(* Logix 5000 project; controller FV vendor 1 type 14 code 217 rev 31.11; software revision 31.00; part 40 of 63 *)
(* tags used below, declared in another part *)
   FV_ALARM : PlantItem;   // ALARM
   FV_ALARM_RawOutput : ALIAS FOR Remote_IO:4:O.Data.5;   // FV_ALARM Audible alarm
   FV_B22 : INT[255];   // YSVFILL_FL YSV filling process flags
   FV_FV25C : PlantItem;   // FV25C
   FV_FV25C_RawOutput : ALIAS FOR Remote_IO:4:O.Data.0;   // FV_FV25C FV 25 cone cooling valve
   FV_FV25J : PlantItem;   // FV25J
   FV_FV25J_RawOutput : ALIAS FOR Remote_IO:4:O.Data.1;   // FV_FV25J FV 25 jacket cooling valve
   FV_FV26C : PlantItem;   // FV26C
   FV_FV26C_RawOutput : ALIAS FOR Remote_IO:9:O.Data.1;   // FV_FV26C FV26 coolant SOV (Cone)
   FV_FV26J : PlantItem;   // FV26J
   FV_FV26J_RawOutput : ALIAS FOR Remote_IO:9:O.Data.0;   // FV_FV26J FV26 coolant SOV (Tank)
   FV_FV27C : PlantItem;   // FV27C
   FV_FV27C_RawOutput : ALIAS FOR Remote_IO:9:O.Data.3;   // FV_FV27C FV27 coolant SOV (Cone)
   FV_FV27J : PlantItem;   // FV27J
   FV_FV27J_RawOutput : ALIAS FOR Remote_IO:9:O.Data.2;   // FV_FV27J FV27 coolant SOV (Tank)
   FV_FV28C : PlantItem;   // FV28C
   FV_FV28C_RawOutput : ALIAS FOR Remote_IO:9:O.Data.5;   // FV_FV28C FV28 coolant SOV (Cone)
   FV_FV28J : PlantItem;   // FV28J
   FV_FV28J_RawOutput : ALIAS FOR Remote_IO:9:O.Data.4;   // FV_FV28J FV28 coolant SOV (Tank)
   FV_FV29C : PlantItem;   // FV29C
   FV_FV29C_RawOutput : ALIAS FOR Remote_IO:9:O.Data.7;   // FV_FV29C FV29 coolant SOV (Cone)
   FV_FV29J : PlantItem;   // FV29J
   FV_FV29J_RawOutput : ALIAS FOR Remote_IO:9:O.Data.6;   // FV_FV29J FV29 coolant SOV (Tank)
   FV_FV30C : PlantItem;   // FV30C
   FV_FV30C_RawOutput : ALIAS FOR Remote_IO:9:O.Data.9;   // FV_FV30C FV30 coolant SOV (Cone)
   FV_FV30J : PlantItem;   // FV30J
   FV_FV30J_RawOutput : ALIAS FOR Remote_IO:9:O.Data.8;   // FV_FV30J FV30 coolant SOV (Tank)
   FV_FV31C : PlantItem;   // FV31C
   FV_FV31C_RawOutput : ALIAS FOR Remote_IO:9:O.Data.11;   // FV_FV31C FV31 coolant SOV (Cone)
   FV_FV31J : PlantItem;   // FV31J
   FV_FV31J_RawOutput : ALIAS FOR Remote_IO:9:O.Data.10;   // FV_FV31J FV31 coolant SOV (Tank)
   FV_N141 : INT[255];   // YSV1 DATA
   FV_N142 : INT[255];   // YSV2 DATA
   FV_N143 : INT[255];   // YSV3 DATA
   FV_N20 : INT[255];   // YSVFILL<PC YSV Filling data fro m PC
   FV_N21 : INT[255];   // YSVFILL>PC YSV Filling process data to PC and contr ol regs
   FV_PUMP1 : PlantItem;   // PUMP1
   FV_PUMP1_RawOutput : ALIAS FOR Remote_IO:4:O.Data.13;   // FV_PUMP1 Coolant recirc.valve 1
   FV_PUMP2 : PlantItem;   // PUMP2
   FV_PUMP2_RawOutput : ALIAS FOR Remote_IO:4:O.Data.14;   // FV_PUMP2 Coolant recirc.valve 2
   FV_PUMP3 : PlantItem;   // PUMP3
   FV_PUMP3_RawOutput : ALIAS FOR Remote_IO:4:O.Data.15;   // FV_PUMP3 Coolant recirc.valve 3
   FV_SOV1 : PlantItem;   // SOV1
   FV_SOV1_RawOutput : ALIAS FOR Remote_IO:5:O.Data.6;   // FV_SOV1 Air supply to reseed pump
   FV_SOV2 : PlantItem;   // SOV2
   FV_SOV2_RawOutput : ALIAS FOR Remote_IO:5:O.Data.7;   // FV_SOV2 Air supply to reseed pump
   FV_T23 : TIMER[10];
   FV_YSV1CV : PlantItem;   // YSV1CV
   FV_YSV1CV_RawOutput : ALIAS FOR Remote_IO:5:O.Data.12;   // FV_YSV1CV
   FV_YSV1J : PlantItem;   // YSV1J
   FV_YSV1J_RawOutput : ALIAS FOR Remote_IO:4:O.Data.9;   // FV_YSV1J YSV 1 cooling valve
   FV_YSV2CV : PlantItem;   // YSV2CV
   FV_YSV2CV_RawOutput : ALIAS FOR Remote_IO:5:O.Data.13;   // FV_YSV2CV
   FV_YSV2J : PlantItem;   // YSV2J
   FV_YSV2J_RawOutput : ALIAS FOR Remote_IO:4:O.Data.11;   // FV_YSV2J YSV 2 cooling valve
   FV_YSV2O : PlantItem;   // YSV2O
   FV_YSV2O_RawOutput : ALIAS FOR Remote_IO:4:O.Data.4;   // FV_YSV2O YSV 2 outlet valve
   FV_YSV2R : PlantItem;   // YSV2R
   FV_YSV2R_RawOutput : ALIAS FOR Remote_IO:4:O.Data.12;   // FV_YSV2R YSV 2 rouser
   FV_YSV3J : PlantItem;   // YSV3J
   FV_YSV3J_RawOutput : ALIAS FOR Remote_IO:4:O.Data.7;   // FV_YSV3J YSV 3 cooling valve
   FV_YSV3O : PlantItem;   // YSV3O
   FV_YSV3O_RawOutput : ALIAS FOR Remote_IO:4:O.Data.6;   // FV_YSV3O YSV 3 outlet valve
   FV_YSV3R : PlantItem;   // YSV3R
   FV_YSV3R_RawOutput : ALIAS FOR Remote_IO:4:O.Data.8;   // FV_YSV3R YSV 3 rouser
(* FV_Common, continued *)

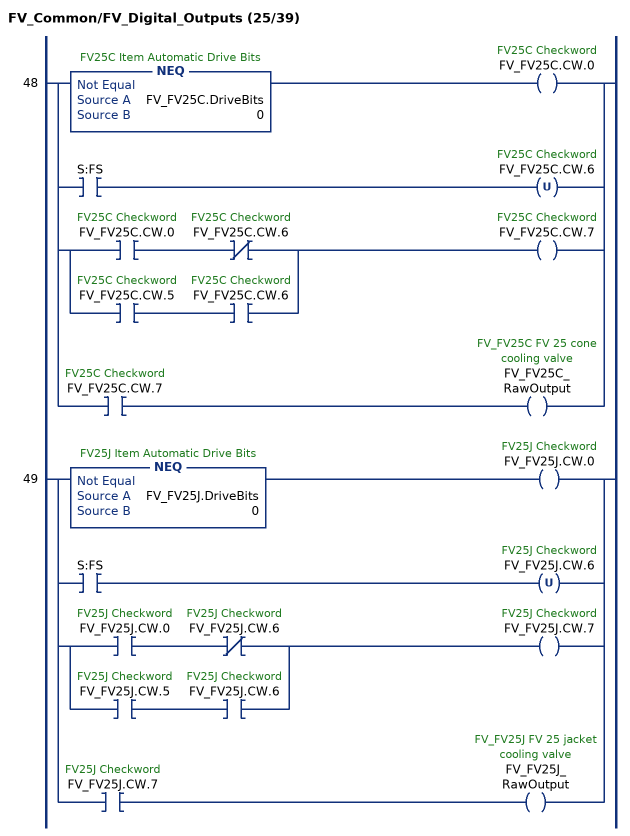
   [picture p849: FV_Common/FV_Digital_Outputs rungs 48-49]
   48: [NEQ(FV_FV25C.DriveBits,0) OTE(FV_FV25C.CW.0) ,XIC(S:FS) OTU(FV_FV25C.CW.6) ,[XIC(FV_FV25C.CW.0) XIO(FV_FV25C.CW.6) ,XIC(FV_FV25C.CW.5) XIC(FV_FV25C.CW.6) ] OTE(FV_FV25C.CW.7) ,XIC(FV_FV25C.CW.7) OTE(FV_FV25C_RawOutput) ];
   49: [NEQ(FV_FV25J.DriveBits,0) OTE(FV_FV25J.CW.0) ,XIC(S:FS) OTU(FV_FV25J.CW.6) ,[XIC(FV_FV25J.CW.0) XIO(FV_FV25J.CW.6) ,XIC(FV_FV25J.CW.5) XIC(FV_FV25J.CW.6) ] OTE(FV_FV25J.CW.7) ,XIC(FV_FV25J.CW.7) OTE(FV_FV25J_RawOutput) ];
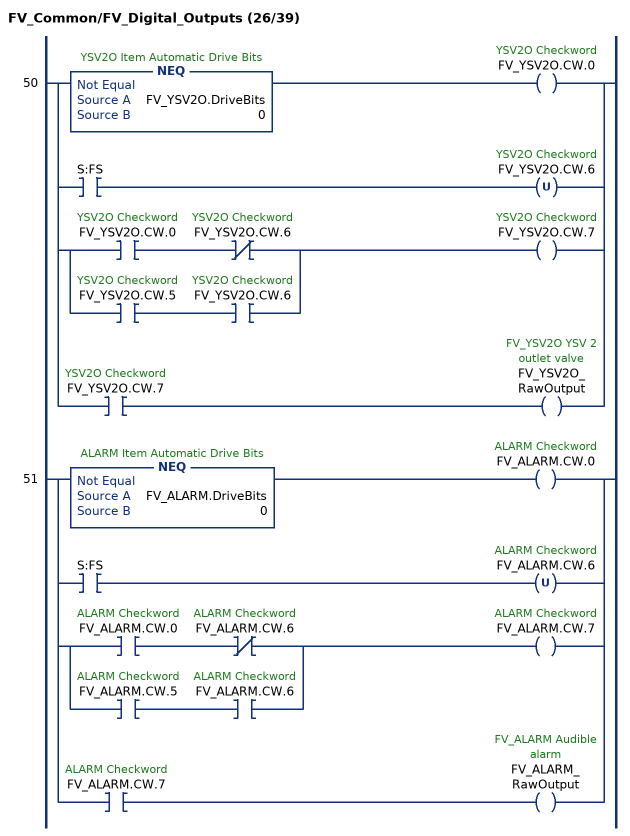
   50: [NEQ(FV_YSV2O.DriveBits,0) OTE(FV_YSV2O.CW.0) ,XIC(S:FS) OTU(FV_YSV2O.CW.6) ,[XIC(FV_YSV2O.CW.0) XIO(FV_YSV2O.CW.6) ,XIC(FV_YSV2O.CW.5) XIC(FV_YSV2O.CW.6) ] OTE(FV_YSV2O.CW.7) ,XIC(FV_YSV2O.CW.7) OTE(FV_YSV2O_RawOutput) ];
   51: [NEQ(FV_ALARM.DriveBits,0) OTE(FV_ALARM.CW.0) ,XIC(S:FS) OTU(FV_ALARM.CW.6) ,[XIC(FV_ALARM.CW.0) XIO(FV_ALARM.CW.6) ,XIC(FV_ALARM.CW.5) XIC(FV_ALARM.CW.6) ] OTE(FV_ALARM.CW.7) ,XIC(FV_ALARM.CW.7) OTE(FV_ALARM_RawOutput) ];
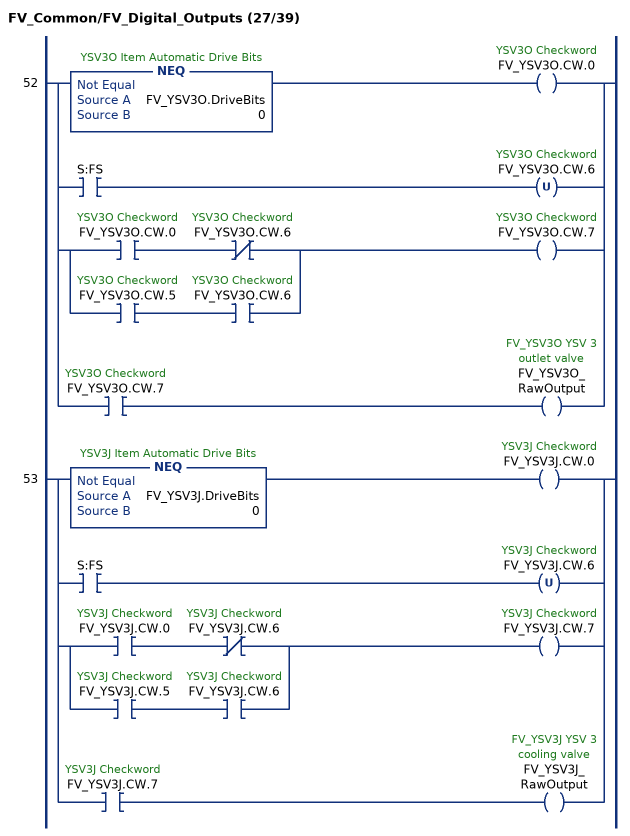
   52: [NEQ(FV_YSV3O.DriveBits,0) OTE(FV_YSV3O.CW.0) ,XIC(S:FS) OTU(FV_YSV3O.CW.6) ,[XIC(FV_YSV3O.CW.0) XIO(FV_YSV3O.CW.6) ,XIC(FV_YSV3O.CW.5) XIC(FV_YSV3O.CW.6) ] OTE(FV_YSV3O.CW.7) ,XIC(FV_YSV3O.CW.7) OTE(FV_YSV3O_RawOutput) ];
   53: [NEQ(FV_YSV3J.DriveBits,0) OTE(FV_YSV3J.CW.0) ,XIC(S:FS) OTU(FV_YSV3J.CW.6) ,[XIC(FV_YSV3J.CW.0) XIO(FV_YSV3J.CW.6) ,XIC(FV_YSV3J.CW.5) XIC(FV_YSV3J.CW.6) ] OTE(FV_YSV3J.CW.7) ,XIC(FV_YSV3J.CW.7) OTE(FV_YSV3J_RawOutput) ];
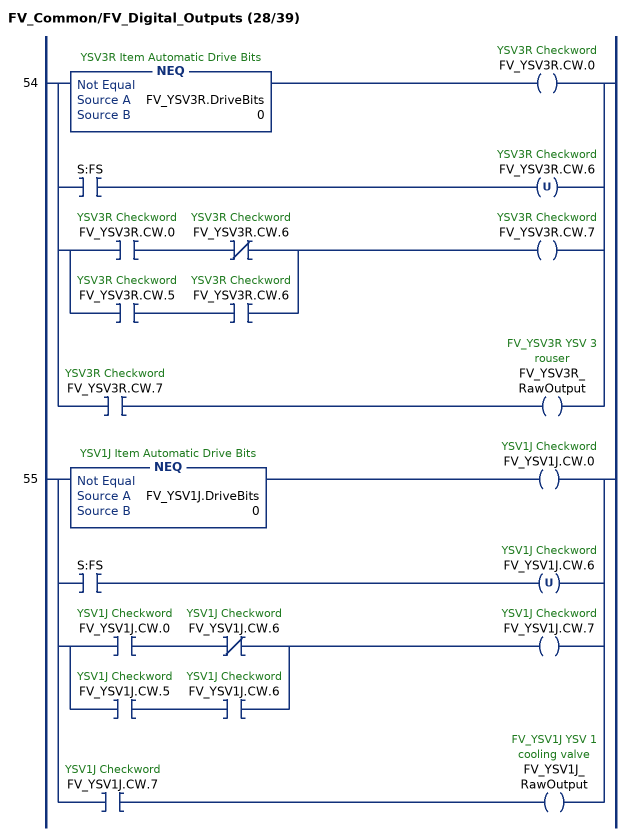
   54: [NEQ(FV_YSV3R.DriveBits,0) OTE(FV_YSV3R.CW.0) ,XIC(S:FS) OTU(FV_YSV3R.CW.6) ,[XIC(FV_YSV3R.CW.0) XIO(FV_YSV3R.CW.6) ,XIC(FV_YSV3R.CW.5) XIC(FV_YSV3R.CW.6) ] OTE(FV_YSV3R.CW.7) ,XIC(FV_YSV3R.CW.7) OTE(FV_YSV3R_RawOutput) ];
   55: [NEQ(FV_YSV1J.DriveBits,0) OTE(FV_YSV1J.CW.0) ,XIC(S:FS) OTU(FV_YSV1J.CW.6) ,[XIC(FV_YSV1J.CW.0) XIO(FV_YSV1J.CW.6) ,XIC(FV_YSV1J.CW.5) XIC(FV_YSV1J.CW.6) ] OTE(FV_YSV1J.CW.7) ,XIC(FV_YSV1J.CW.7) OTE(FV_YSV1J_RawOutput) ];
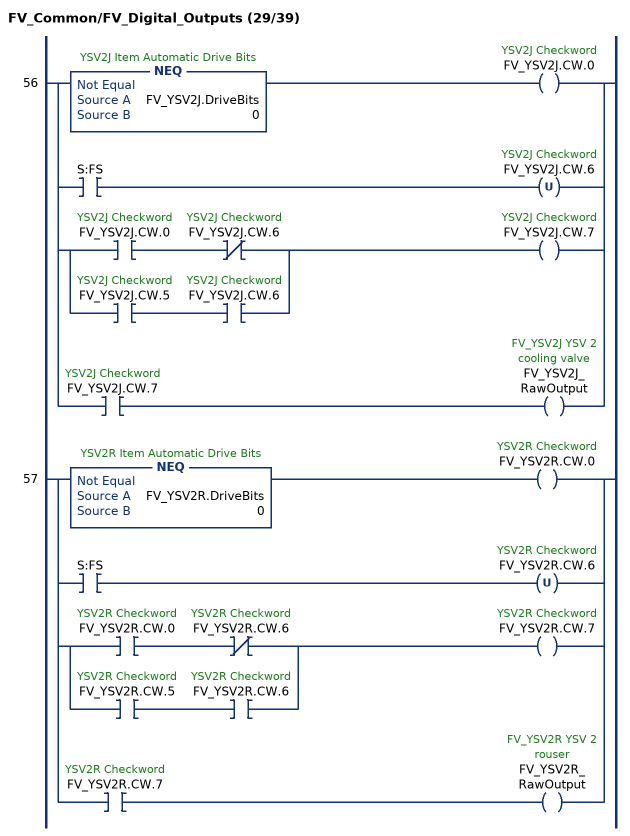
   56: [NEQ(FV_YSV2J.DriveBits,0) OTE(FV_YSV2J.CW.0) ,XIC(S:FS) OTU(FV_YSV2J.CW.6) ,[XIC(FV_YSV2J.CW.0) XIO(FV_YSV2J.CW.6) ,XIC(FV_YSV2J.CW.5) XIC(FV_YSV2J.CW.6) ] OTE(FV_YSV2J.CW.7) ,XIC(FV_YSV2J.CW.7) OTE(FV_YSV2J_RawOutput) ];
   57: [NEQ(FV_YSV2R.DriveBits,0) OTE(FV_YSV2R.CW.0) ,XIC(S:FS) OTU(FV_YSV2R.CW.6) ,[XIC(FV_YSV2R.CW.0) XIO(FV_YSV2R.CW.6) ,XIC(FV_YSV2R.CW.5) XIC(FV_YSV2R.CW.6) ] OTE(FV_YSV2R.CW.7) ,XIC(FV_YSV2R.CW.7) OTE(FV_YSV2R_RawOutput) ];
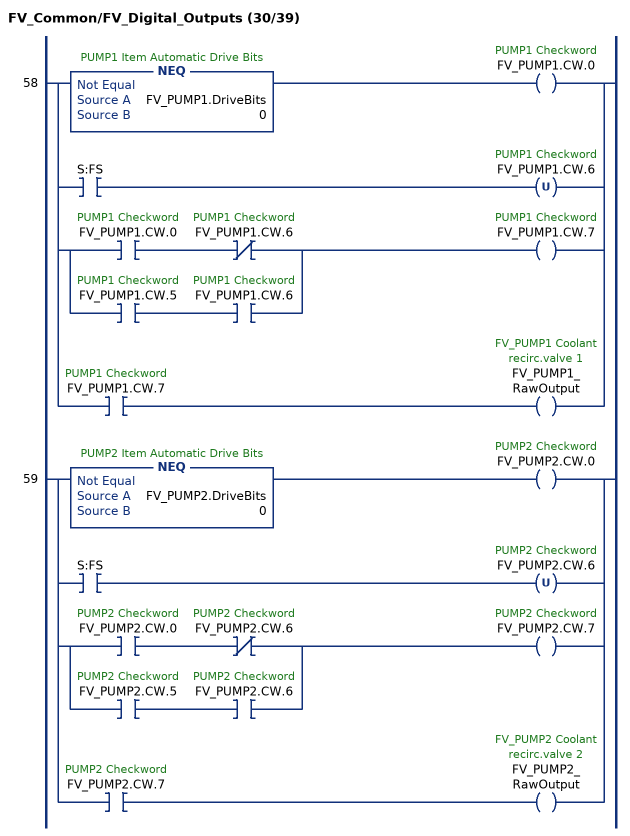
   58: [NEQ(FV_PUMP1.DriveBits,0) OTE(FV_PUMP1.CW.0) ,XIC(S:FS) OTU(FV_PUMP1.CW.6) ,[XIC(FV_PUMP1.CW.0) XIO(FV_PUMP1.CW.6) ,XIC(FV_PUMP1.CW.5) XIC(FV_PUMP1.CW.6) ] OTE(FV_PUMP1.CW.7) ,XIC(FV_PUMP1.CW.7) OTE(FV_PUMP1_RawOutput) ];
   59: [NEQ(FV_PUMP2.DriveBits,0) OTE(FV_PUMP2.CW.0) ,XIC(S:FS) OTU(FV_PUMP2.CW.6) ,[XIC(FV_PUMP2.CW.0) XIO(FV_PUMP2.CW.6) ,XIC(FV_PUMP2.CW.5) XIC(FV_PUMP2.CW.6) ] OTE(FV_PUMP2.CW.7) ,XIC(FV_PUMP2.CW.7) OTE(FV_PUMP2_RawOutput) ];
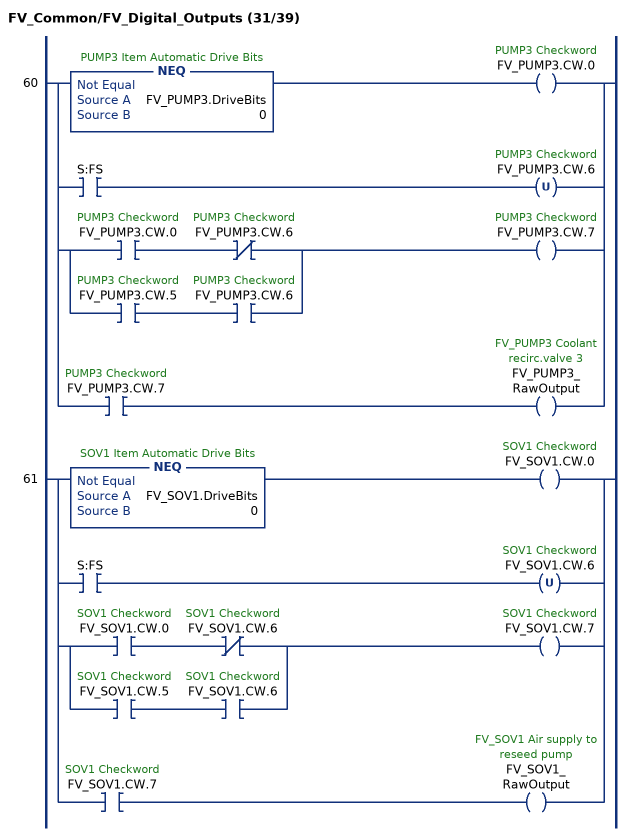
   60: [NEQ(FV_PUMP3.DriveBits,0) OTE(FV_PUMP3.CW.0) ,XIC(S:FS) OTU(FV_PUMP3.CW.6) ,[XIC(FV_PUMP3.CW.0) XIO(FV_PUMP3.CW.6) ,XIC(FV_PUMP3.CW.5) XIC(FV_PUMP3.CW.6) ] OTE(FV_PUMP3.CW.7) ,XIC(FV_PUMP3.CW.7) OTE(FV_PUMP3_RawOutput) ];
   61: [NEQ(FV_SOV1.DriveBits,0) OTE(FV_SOV1.CW.0) ,XIC(S:FS) OTU(FV_SOV1.CW.6) ,[XIC(FV_SOV1.CW.0) XIO(FV_SOV1.CW.6) ,XIC(FV_SOV1.CW.5) XIC(FV_SOV1.CW.6) ] OTE(FV_SOV1.CW.7) ,XIC(FV_SOV1.CW.7) OTE(FV_SOV1_RawOutput) ];
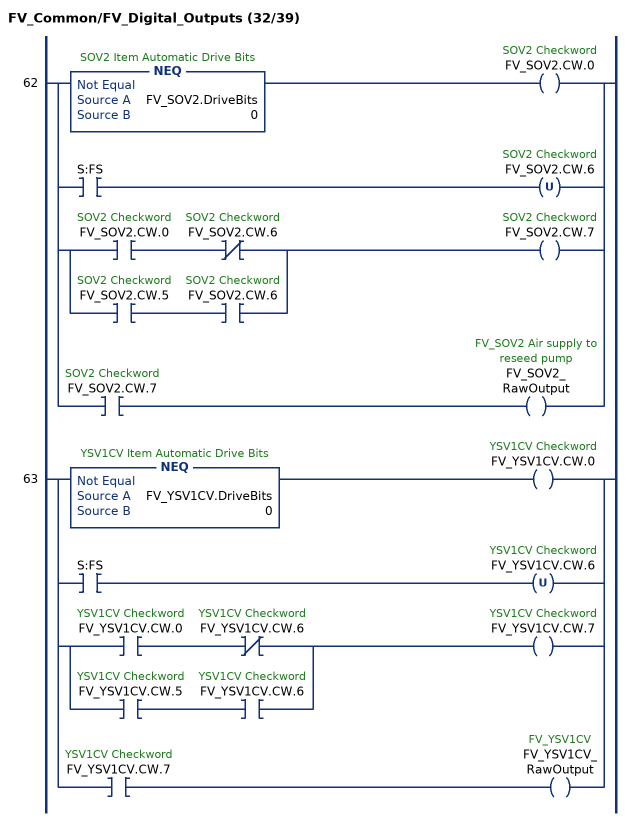
   62: [NEQ(FV_SOV2.DriveBits,0) OTE(FV_SOV2.CW.0) ,XIC(S:FS) OTU(FV_SOV2.CW.6) ,[XIC(FV_SOV2.CW.0) XIO(FV_SOV2.CW.6) ,XIC(FV_SOV2.CW.5) XIC(FV_SOV2.CW.6) ] OTE(FV_SOV2.CW.7) ,XIC(FV_SOV2.CW.7) OTE(FV_SOV2_RawOutput) ];
   63: [NEQ(FV_YSV1CV.DriveBits,0) OTE(FV_YSV1CV.CW.0) ,XIC(S:FS) OTU(FV_YSV1CV.CW.6) ,[XIC(FV_YSV1CV.CW.0) XIO(FV_YSV1CV.CW.6) ,XIC(FV_YSV1CV.CW.5) XIC(FV_YSV1CV.CW.6) ] OTE(FV_YSV1CV.CW.7) ,XIC(FV_YSV1CV.CW.7) OTE(FV_YSV1CV_RawOutput) ];
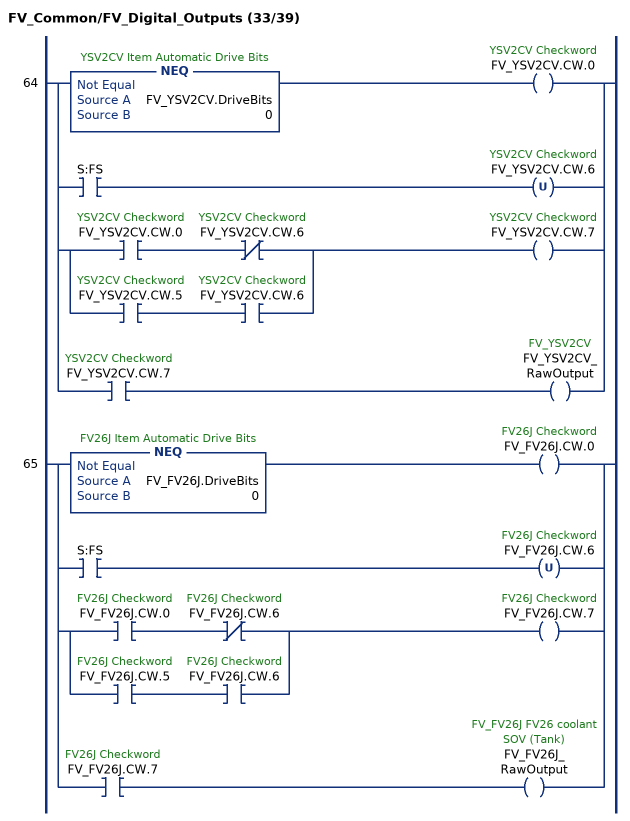
   64: [NEQ(FV_YSV2CV.DriveBits,0) OTE(FV_YSV2CV.CW.0) ,XIC(S:FS) OTU(FV_YSV2CV.CW.6) ,[XIC(FV_YSV2CV.CW.0) XIO(FV_YSV2CV.CW.6) ,XIC(FV_YSV2CV.CW.5) XIC(FV_YSV2CV.CW.6) ] OTE(FV_YSV2CV.CW.7) ,XIC(FV_YSV2CV.CW.7) OTE(FV_YSV2CV_RawOutput) ];
   65: [NEQ(FV_FV26J.DriveBits,0) OTE(FV_FV26J.CW.0) ,XIC(S:FS) OTU(FV_FV26J.CW.6) ,[XIC(FV_FV26J.CW.0) XIO(FV_FV26J.CW.6) ,XIC(FV_FV26J.CW.5) XIC(FV_FV26J.CW.6) ] OTE(FV_FV26J.CW.7) ,XIC(FV_FV26J.CW.7) OTE(FV_FV26J_RawOutput) ];
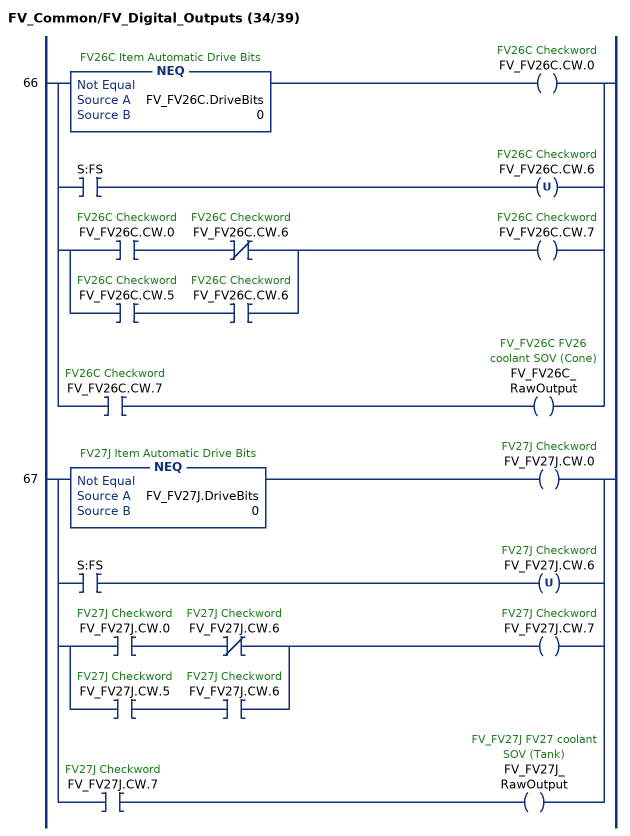
   66: [NEQ(FV_FV26C.DriveBits,0) OTE(FV_FV26C.CW.0) ,XIC(S:FS) OTU(FV_FV26C.CW.6) ,[XIC(FV_FV26C.CW.0) XIO(FV_FV26C.CW.6) ,XIC(FV_FV26C.CW.5) XIC(FV_FV26C.CW.6) ] OTE(FV_FV26C.CW.7) ,XIC(FV_FV26C.CW.7) OTE(FV_FV26C_RawOutput) ];
   67: [NEQ(FV_FV27J.DriveBits,0) OTE(FV_FV27J.CW.0) ,XIC(S:FS) OTU(FV_FV27J.CW.6) ,[XIC(FV_FV27J.CW.0) XIO(FV_FV27J.CW.6) ,XIC(FV_FV27J.CW.5) XIC(FV_FV27J.CW.6) ] OTE(FV_FV27J.CW.7) ,XIC(FV_FV27J.CW.7) OTE(FV_FV27J_RawOutput) ];
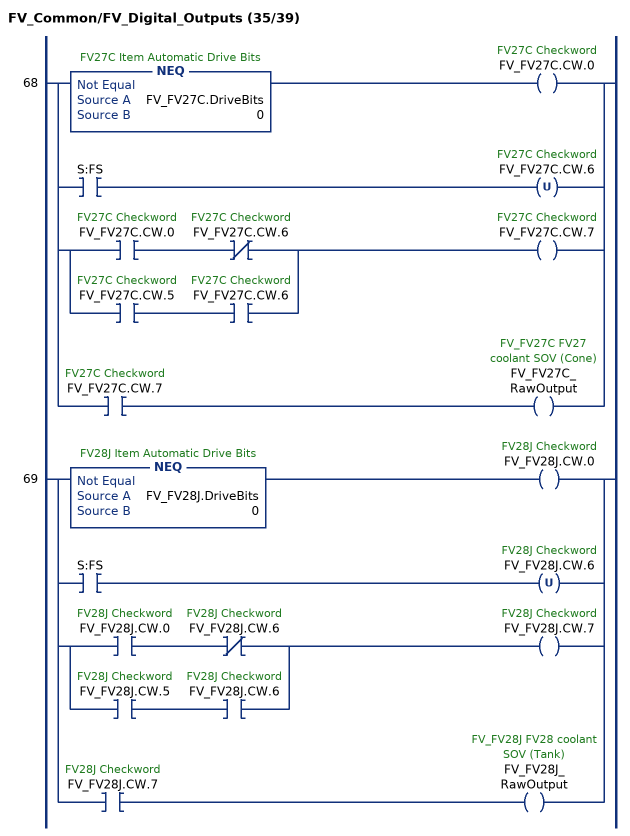
   68: [NEQ(FV_FV27C.DriveBits,0) OTE(FV_FV27C.CW.0) ,XIC(S:FS) OTU(FV_FV27C.CW.6) ,[XIC(FV_FV27C.CW.0) XIO(FV_FV27C.CW.6) ,XIC(FV_FV27C.CW.5) XIC(FV_FV27C.CW.6) ] OTE(FV_FV27C.CW.7) ,XIC(FV_FV27C.CW.7) OTE(FV_FV27C_RawOutput) ];
   69: [NEQ(FV_FV28J.DriveBits,0) OTE(FV_FV28J.CW.0) ,XIC(S:FS) OTU(FV_FV28J.CW.6) ,[XIC(FV_FV28J.CW.0) XIO(FV_FV28J.CW.6) ,XIC(FV_FV28J.CW.5) XIC(FV_FV28J.CW.6) ] OTE(FV_FV28J.CW.7) ,XIC(FV_FV28J.CW.7) OTE(FV_FV28J_RawOutput) ];
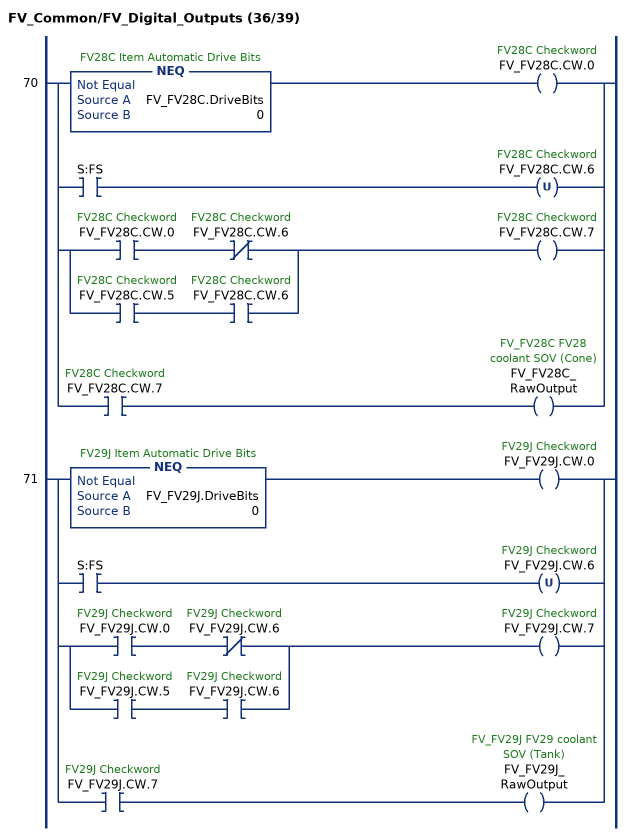
   70: [NEQ(FV_FV28C.DriveBits,0) OTE(FV_FV28C.CW.0) ,XIC(S:FS) OTU(FV_FV28C.CW.6) ,[XIC(FV_FV28C.CW.0) XIO(FV_FV28C.CW.6) ,XIC(FV_FV28C.CW.5) XIC(FV_FV28C.CW.6) ] OTE(FV_FV28C.CW.7) ,XIC(FV_FV28C.CW.7) OTE(FV_FV28C_RawOutput) ];
   71: [NEQ(FV_FV29J.DriveBits,0) OTE(FV_FV29J.CW.0) ,XIC(S:FS) OTU(FV_FV29J.CW.6) ,[XIC(FV_FV29J.CW.0) XIO(FV_FV29J.CW.6) ,XIC(FV_FV29J.CW.5) XIC(FV_FV29J.CW.6) ] OTE(FV_FV29J.CW.7) ,XIC(FV_FV29J.CW.7) OTE(FV_FV29J_RawOutput) ];
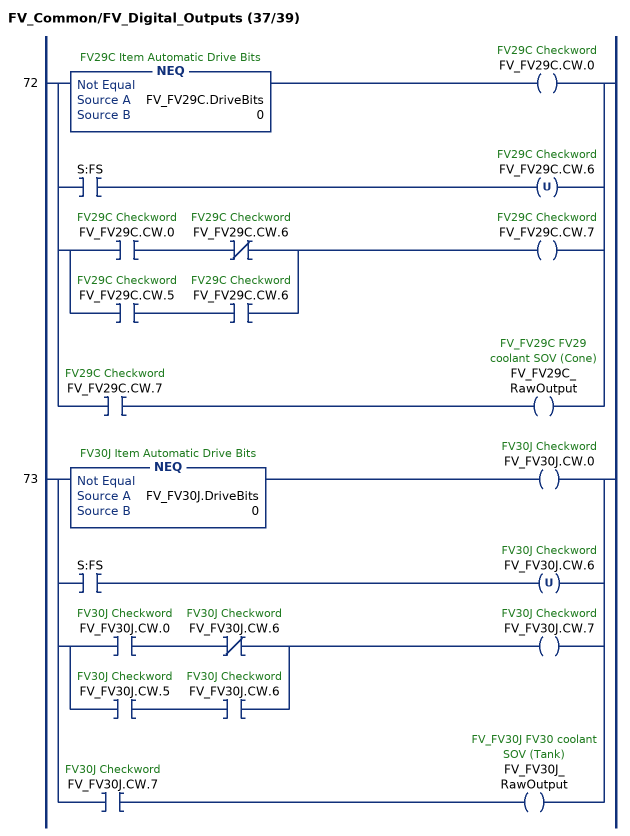
   72: [NEQ(FV_FV29C.DriveBits,0) OTE(FV_FV29C.CW.0) ,XIC(S:FS) OTU(FV_FV29C.CW.6) ,[XIC(FV_FV29C.CW.0) XIO(FV_FV29C.CW.6) ,XIC(FV_FV29C.CW.5) XIC(FV_FV29C.CW.6) ] OTE(FV_FV29C.CW.7) ,XIC(FV_FV29C.CW.7) OTE(FV_FV29C_RawOutput) ];
   73: [NEQ(FV_FV30J.DriveBits,0) OTE(FV_FV30J.CW.0) ,XIC(S:FS) OTU(FV_FV30J.CW.6) ,[XIC(FV_FV30J.CW.0) XIO(FV_FV30J.CW.6) ,XIC(FV_FV30J.CW.5) XIC(FV_FV30J.CW.6) ] OTE(FV_FV30J.CW.7) ,XIC(FV_FV30J.CW.7) OTE(FV_FV30J_RawOutput) ];
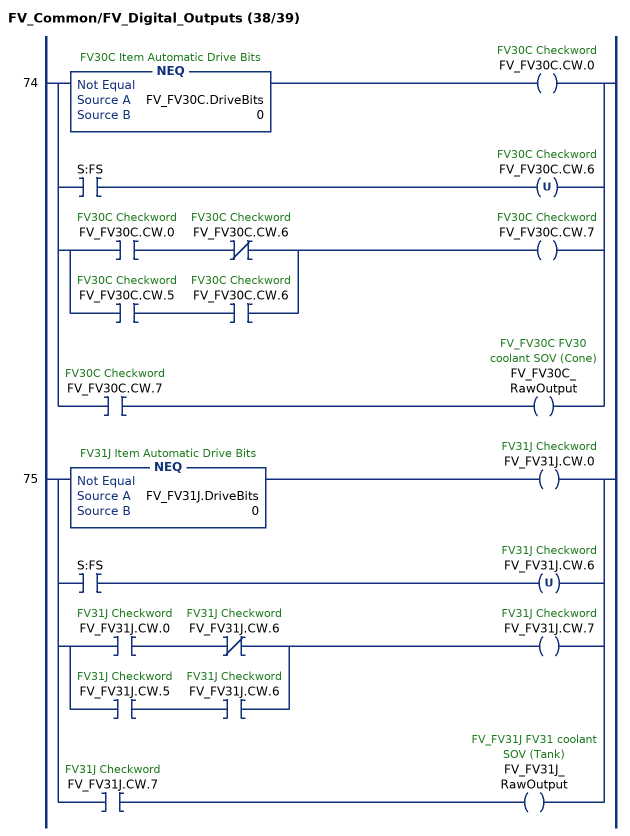
   74: [NEQ(FV_FV30C.DriveBits,0) OTE(FV_FV30C.CW.0) ,XIC(S:FS) OTU(FV_FV30C.CW.6) ,[XIC(FV_FV30C.CW.0) XIO(FV_FV30C.CW.6) ,XIC(FV_FV30C.CW.5) XIC(FV_FV30C.CW.6) ] OTE(FV_FV30C.CW.7) ,XIC(FV_FV30C.CW.7) OTE(FV_FV30C_RawOutput) ];
   75: [NEQ(FV_FV31J.DriveBits,0) OTE(FV_FV31J.CW.0) ,XIC(S:FS) OTU(FV_FV31J.CW.6) ,[XIC(FV_FV31J.CW.0) XIO(FV_FV31J.CW.6) ,XIC(FV_FV31J.CW.5) XIC(FV_FV31J.CW.6) ] OTE(FV_FV31J.CW.7) ,XIC(FV_FV31J.CW.7) OTE(FV_FV31J_RawOutput) ];
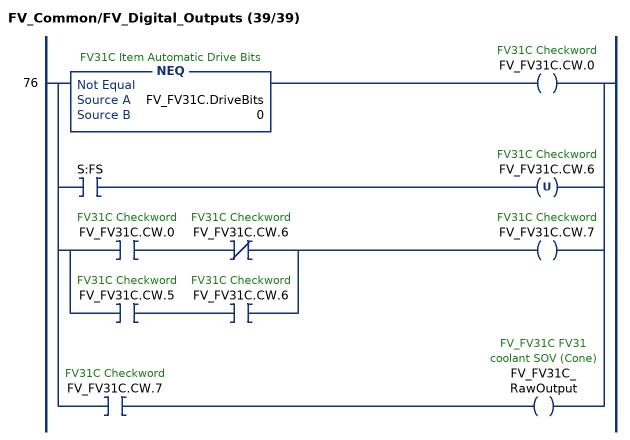
   76: [NEQ(FV_FV31C.DriveBits,0) OTE(FV_FV31C.CW.0) ,XIC(S:FS) OTU(FV_FV31C.CW.6) ,[XIC(FV_FV31C.CW.0) XIO(FV_FV31C.CW.6) ,XIC(FV_FV31C.CW.5) XIC(FV_FV31C.CW.6) ] OTE(FV_FV31C.CW.7) ,XIC(FV_FV31C.CW.7) OTE(FV_FV31C_RawOutput) ];
END_ROUTINE

ROUTINE FV_FILLYSV_CP_11   (* ladder *)
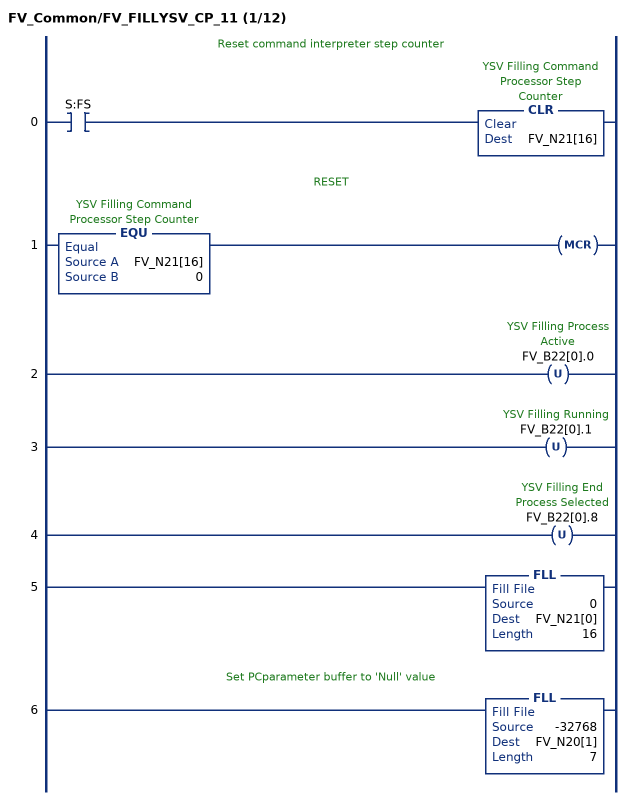
   // Reset command interpreter step counter
   0: XIC(S:FS)CLR(FV_N21[16]);
   // RESET
   1: EQU(FV_N21[16],0)MCR();
   2: OTU(FV_B22[0].0);
   3: OTU(FV_B22[0].1);
   4: OTU(FV_B22[0].8);
   5: FLL(0,FV_N21[0],16);
   // Set PCparameter buffer to 'Null' value
   6: FLL(-32768,FV_N20[1],7);
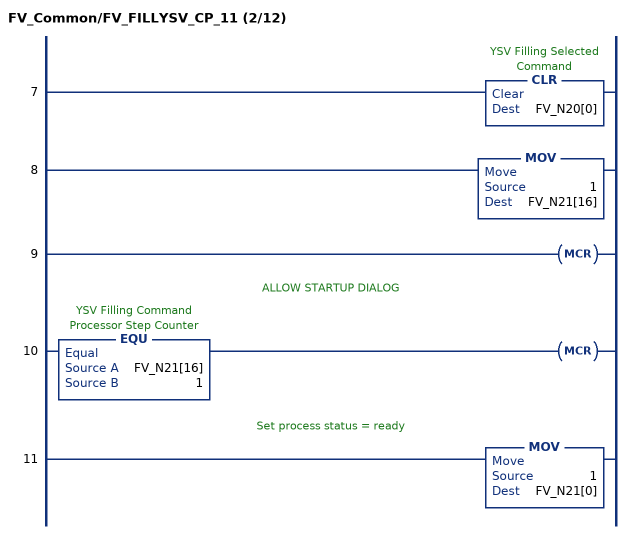
   7: CLR(FV_N20[0]);
   8: MOV(1,FV_N21[16]);
   9: MCR();
   // ALLOW STARTUP DIALOG
   10: EQU(FV_N21[16],1)MCR();
   // Set process status = ready
   11: MOV(1,FV_N21[0]);
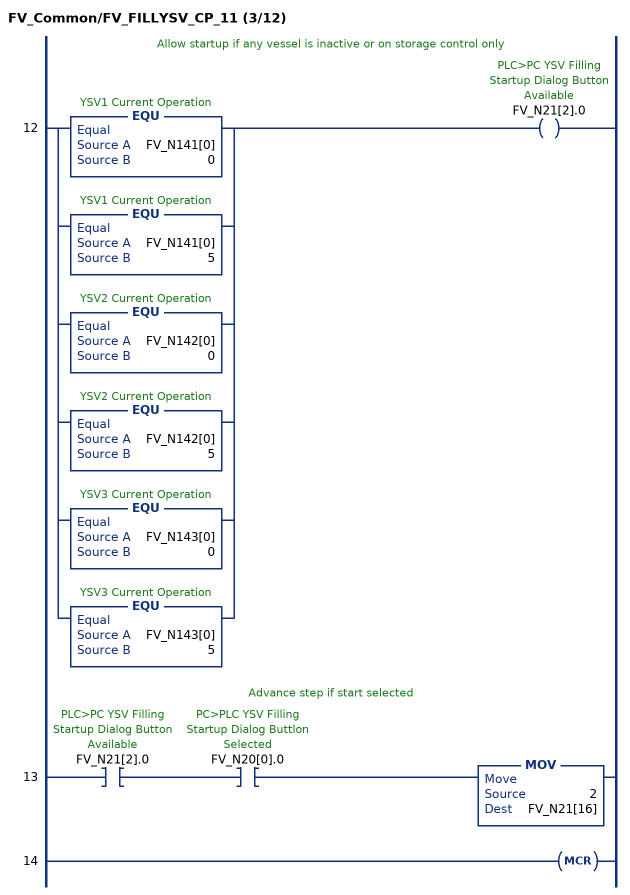
   // Allow startup if any vessel is inactive or on storage control only
   12: [[EQU(FV_N141[0],0) ,EQU(FV_N141[0],5) ] ,[EQU(FV_N142[0],0) ,EQU(FV_N142[0],5) ] ,[EQU(FV_N143[0],0) ,EQU(FV_N143[0],5) ] ]OTE(FV_N21[2].0);
   // Advance step if start selected
   13: XIC(FV_N21[2].0)XIC(FV_N20[0].0)MOV(2,FV_N21[16]);
   14: MCR();
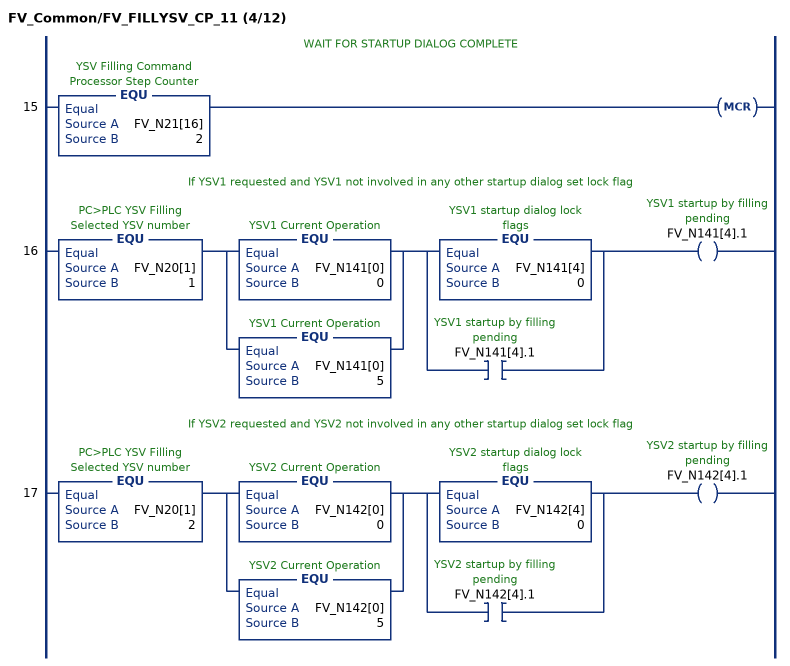
   // WAIT FOR STARTUP DIALOG COMPLETE
   15: EQU(FV_N21[16],2)MCR();
   // If YSV1 requested and YSV1 not involved in any other startup dialog set lock flag
   16: EQU(FV_N20[1],1)[EQU(FV_N141[0],0) ,EQU(FV_N141[0],5) ][EQU(FV_N141[4],0) ,XIC(FV_N141[4].1) ]OTE(FV_N141[4].1);
   // If YSV2 requested and YSV2 not involved in any other startup dialog set lock flag
   17: EQU(FV_N20[1],2)[EQU(FV_N142[0],0) ,EQU(FV_N142[0],5) ][EQU(FV_N142[4],0) ,XIC(FV_N142[4].1) ]OTE(FV_N142[4].1);
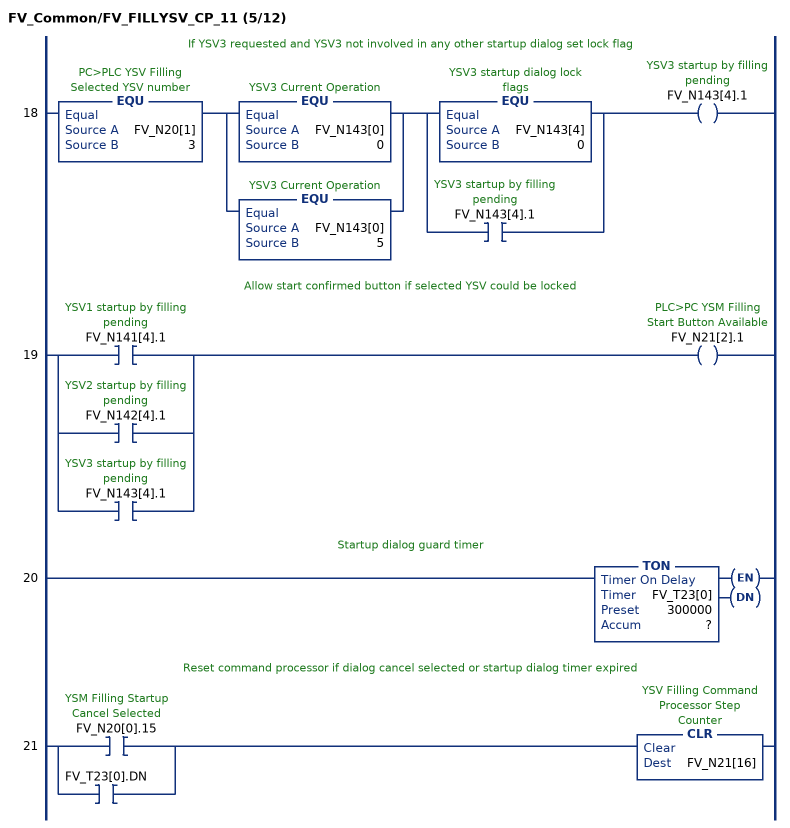
   // If YSV3 requested and YSV3 not involved in any other startup dialog set lock flag
   18: EQU(FV_N20[1],3)[EQU(FV_N143[0],0) ,EQU(FV_N143[0],5) ][EQU(FV_N143[4],0) ,XIC(FV_N143[4].1) ]OTE(FV_N143[4].1);
   // Allow start confirmed button if selected YSV could be locked
   19: [XIC(FV_N141[4].1) ,XIC(FV_N142[4].1) ,XIC(FV_N143[4].1) ]OTE(FV_N21[2].1);
   // Startup dialog guard timer
   20: TON(FV_T23[0],?,?);
   // Reset command processor if dialog cancel selected or startup dialog timer expired
   21: [XIC(FV_N20[0].15) ,XIC(FV_T23[0].DN) ]CLR(FV_N21[16]);
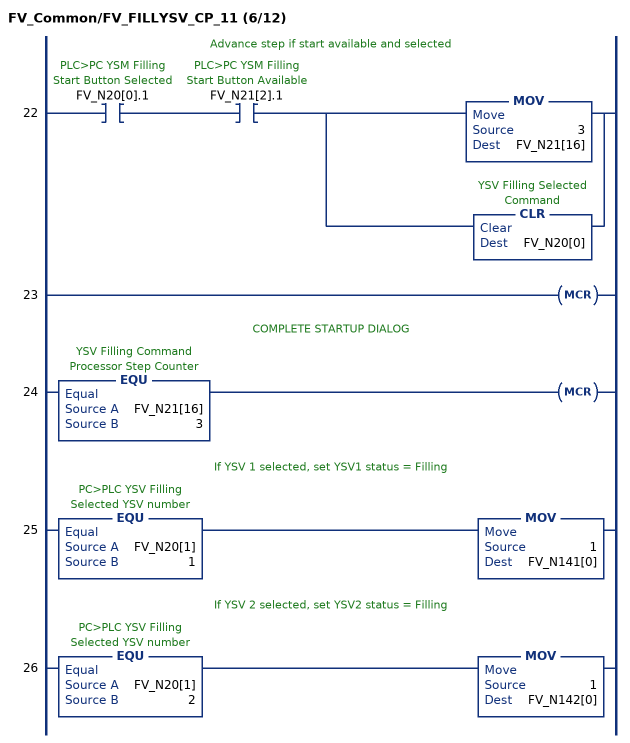
   // Advance step if start available and selected
   22: XIC(FV_N20[0].1)XIC(FV_N21[2].1)[MOV(3,FV_N21[16]) ,CLR(FV_N20[0]) ];
   23: MCR();
   // COMPLETE STARTUP DIALOG
   24: EQU(FV_N21[16],3)MCR();
   // If YSV 1 selected, set YSV1 status = Filling
   25: EQU(FV_N20[1],1)MOV(1,FV_N141[0]);
   // If YSV 2 selected, set YSV2 status = Filling
   26: EQU(FV_N20[1],2)MOV(1,FV_N142[0]);
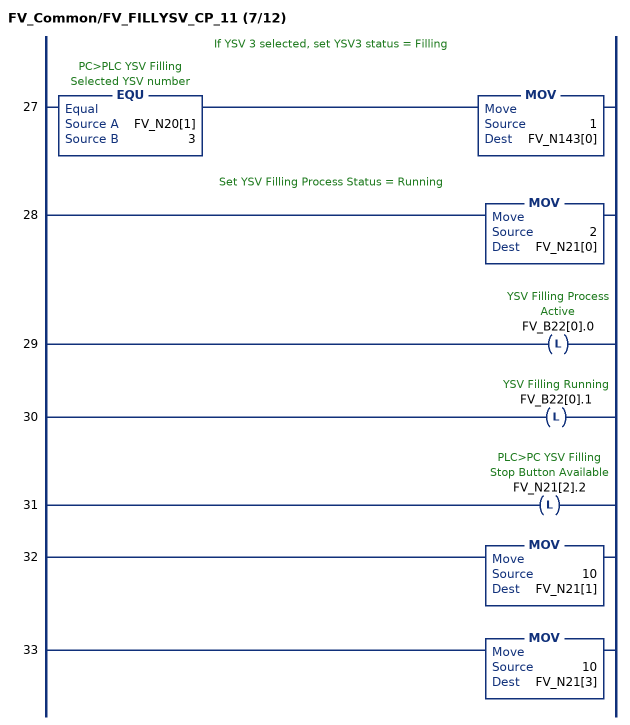
   // If YSV 3 selected, set YSV3 status = Filling
   27: EQU(FV_N20[1],3)MOV(1,FV_N143[0]);
   // Set YSV Filling Process Status = Running
   28: MOV(2,FV_N21[0]);
   29: OTL(FV_B22[0].0);
   30: OTL(FV_B22[0].1);
   31: OTL(FV_N21[2].2);
   32: MOV(10,FV_N21[1]);
   33: MOV(10,FV_N21[3]);
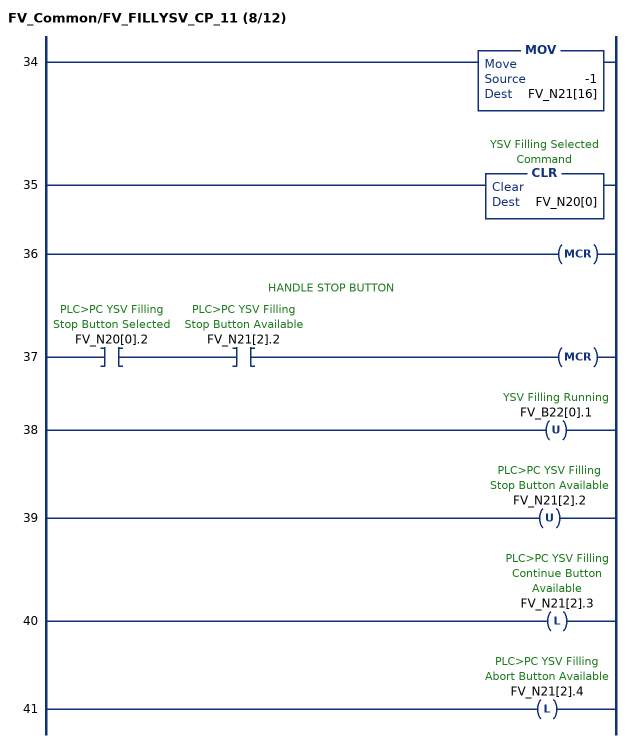
   34: MOV(-1,FV_N21[16]);
   35: CLR(FV_N20[0]);
   36: MCR();
   // HANDLE STOP BUTTON
   37: XIC(FV_N20[0].2)XIC(FV_N21[2].2)MCR();
   38: OTU(FV_B22[0].1);
   39: OTU(FV_N21[2].2);
   40: OTL(FV_N21[2].3);
   41: OTL(FV_N21[2].4);
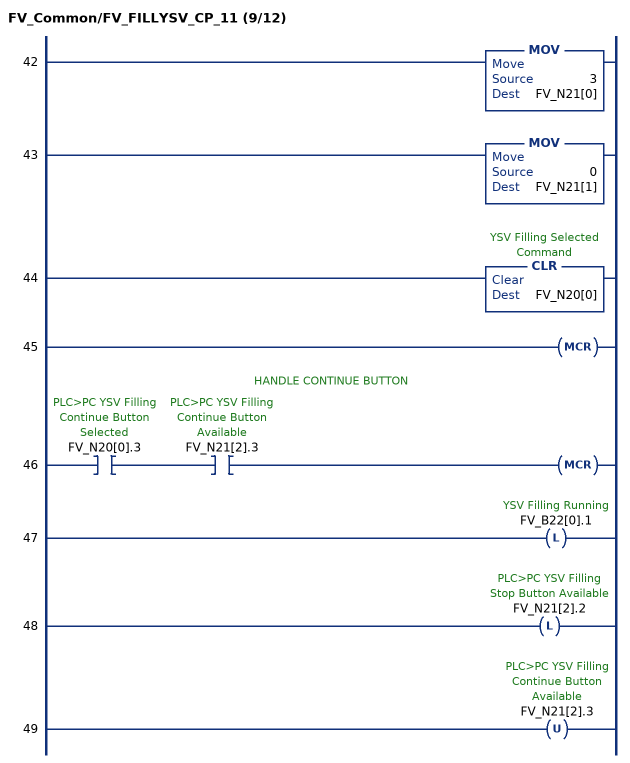
   42: MOV(3,FV_N21[0]);
   43: MOV(0,FV_N21[1]);
   44: CLR(FV_N20[0]);
   45: MCR();
   // HANDLE CONTINUE BUTTON
   46: XIC(FV_N20[0].3)XIC(FV_N21[2].3)MCR();
   47: OTL(FV_B22[0].1);
   48: OTL(FV_N21[2].2);
   49: OTU(FV_N21[2].3);
